// TIA Portal project "TIA_V16_ScalingFunctionExample" (V16)

(* hardware
DEVICE "S71500/ET200MP station_1"  S7-1500 station
   slot 0: "Rail_0"  Rack  6ES7 590-1***0-0AA0
   slot 0: "PS 25W 24VDC_1"  PS 25W 24VDC  6ES7 505-0KA00-0AB0  V1.0
   slot 1: "PLC_1"  CPU 1511F-1 PN  6ES7 511-1FK01-0AB0  V1.8
   slot 2: "DI 16x24VDC HF_1"  DI 16x24VDC HF  6ES7 521-1BH00-0AB0  V2.0
   slot 3: "DQ 16x24VDC/0.5A ST_1"  DQ 16x24VDC/0.5A ST  6ES7 522-1BH00-0AB0  V2.0
   slot 4: "AI 4xU/I/RTD/TC ST_1"  AI 4xU/I/RTD/TC ST  6ES7 531-7QD00-0AB0  V1.0
   slot 5: "AQ 4xU/I ST_1"  AQ 4xU/I ST  6ES7 532-5HD00-0AB0  V2.0
DEVICE "SCALANCE X005"  SCALANCE X-Station
   slot 0: "SCALANCE X rack"  Rail
   slot 0: "Switch_1"  6GK5 005-0BA00-1AA3  V1.0
DEVICE "HMI_1"  TP1200 Comfort
   slot 0: "HMI_1"  TP1200 Comfort  6AV2 124-0MC01-0AX0  16.0.0.0
   slot 1: "HMI_RT_1"  TP1200 Comfort  6AV2 124-0MC01-0AX0  16.0.0.0
   slot 5: "HMI_1.IE_CP_1"  PROFINET Interface  16.0.0.0
      slot 1: "PROFINET Interface_1"  PROFINET Interface
         slot 1: "Port_1"  Port
         slot 2: "Port_2"  Port
   slot 7: "HMI_1.MPI/DP_CP_1"  MPI/DP Interface  16.0.0.0
*)

// ===== PLC "PLC_1"  CPU 1511F-1 PN =====
// protected blocks, not shown: "Main_Safety_RTG1_1", "Main_Safety_RTG1_DB_1"

TYPE "Data Exchange"
TITLE = Data Exchange Between Working Areas
VERSION : 0.1
   STRUCT
      "Working Area 1 Completed" : Bool;
      "Working Area 1 Can Work" : Bool;
      "Working Area 1 Can't Work" : Bool;
      "Working Area 2 Completed" : Bool;
      "Working Area 2 Can Work" : Bool;
      "Working Area 2 Can't  Work" : Bool;
      "Working Area 3 Completed" : Bool;
      "Working Area 3 Can Work" : Bool;
      "Working Area 3 Can't Work" : Bool;
      "Working Area 4 Completed" : Bool;
      "Working Area 4 Can Work" : Bool;
      "Working Area 4 Can't Work" : Bool;
      "WA2 Proof Station OK" : Bool;
      "WA2 Proof Station NOk" : Bool;
      "WA3 Ignition OK" : Bool;
      "WA3 Ignition NOK" : Bool;
      "WA3 Chamber Pressure OK" : Bool;
      "WA3 Chamber Pressure NOK" : Bool;
      Spare1 : Bool;
      Spare2 : Bool;
      Spare3 : Bool;
      Spare4 : Bool;
      Spare5 : Bool;
      Spare6 : Bool;
      Spare7 : Bool;
      Spare8 : Bool;
      Spare9 : Bool;
      Spare10 : Bool;
      Spare11 : Bool;
      Spare12 : Bool;
      Spare13 : Bool;
      Spare14 : Bool;
      Element_1 : Int;
      Element_2 : Int;
      Element_3 : Int;
      Element_4 : Int;
      Element_5 : Int;
      Element_6 : Real;
      Element_8 : Real;
      Element_7 : Real;
      Element_9 : Real;
      Element_10 : Real;
      Rec_PartID : Int;   // Part Record ID Number / 记录ID号
      Rec_Dose_Setting : DInt;   // record recipe dosing setting / 充气设置
      Rec_Gas_Setting_1 : Real;   // record recipe gas setting for shot 1
      Rec_O2_Setting_1 : Real;   // record recipe O2 setting for shot 2
      Rec_Part_Qty : Int;   // record part fixture quanity / 夹具数量
      Rec_Part_weight : Real;   // record recipe part weight
      Rec_shot_type : Int;   // Record recipe shot type
      Rec_Part_image : Array[1..14] of Char;   // PLC part image
      Rec_Fixture_Ref : Array[1..14] of Char;   // record part fixture reference / 夹具参考
      Rec_Part_material : Array[1..14] of Char;   // record part material / 零件材料
      Rec_Part_Name : Array[1..14] of Char;   // record name of part / 记录名称
      Rec_Part_Ref : String[14] := '0';   // record part reference / 零件参考
      Rec_Mix_type1 : Bool;   // record recipe mix type
      Rec_Gas_Setting_2 : Real;   // record recipe gas setting for shot 2
      Rec_O2_Setting_2 : Real;   // record recipe O2 setting for shot 2
      Val_Calibrated_Gas : Int;
      Val_Calibrated_O2 : Int;
      Val_Cailbrated_Gas_Upper : Int;
      Val_Calibrated_Gas_Lower : Int;
      Val_Calibrated_O2_Upper : Int;
      Val_Calibrated_O2_Lower : Int;
      Val_Setting_Gas_Shot_1 : Int;   // Value sent to analog controller for output / 输出值
      Val_Setting_Gas_Shot_2 : Int;   // Value sent to analog controller for output / 输出值
      Val_Setting_O2_Shot_1 : Int := 750;   // Value sent to analog controller for output / 输出值
      Val_Setting_O2_Shot_2 : Int;   // Value sent to analog controller for output / 输出值
      Dose_Setting_Applied : DInt;   // Dosing Stroke Value Applied to Cycle
      BAR_CODE : String[20];
      Rec_MFC_Gas_Setpoint : DInt;
      Rec_MFC_O2_Setpoint : DInt;
   END_STRUCT;
   // Rec_Part_image[1] := '0';
   // Rec_Fixture_Ref[1] := '0';
   // Rec_Part_material[1] := '0';
   // Rec_Part_Name[1] := '0';
END_TYPE

TYPE "UDT_ScalingInputOutput"
   STRUCT
      IN_PV : Word;   // input process value
      IN_OUT_VAL_MIN : Real;   // output value Low limit
      IN_OUT_VAL_MAX : Real;   // output value High limit
      IN_MIN : Real;   // input value Low limit
      IN_MAX : Real;   // input value High limit
      OUT_VAL : Real;   // Output scaled signal
   END_STRUCT;
END_TYPE

TYPE "UDT_ValveActiveConditions_Type_A001"
   STRUCT
      ConditionA : Bool;
      ConditionB : Bool;
      ConditionC : Bool;
   END_STRUCT;
END_TYPE

TYPE "UDT_ValveActiveConditions_Type_A002"
   STRUCT
      ConditionA : Bool;
      ConditionB : Bool;
   END_STRUCT;
END_TYPE

TYPE "UDT_ScalingInput"
   STRUCT
      IN_PV : Word;   // input process value
      IN_OUT_VAL_MIN : Real;   // output value Low limit
      IN_OUT_VAL_MAX : Real;   // output value High limit
      IN_MIN : Real;   // input value Low limit
      IN_MAX : Real;   // input value High limit
   END_STRUCT;
END_TYPE

TYPE "UDT_ScalingOutput"
   STRUCT
      OUT_VAL : Real;   // Output scaled signal
   END_STRUCT;
END_TYPE

// folder: 101_Group_01

DATA_BLOCK "101_DB_ValvesControl"   // DB101
TITLE = 101_DB_Calc_WarmUp_Dosing
{ S7_Optimized_Access := 'FALSE' }
AUTHOR : Jamal
VERSION : 0.1
   VAR
      Valve_1001_Inputs : "UDT_ScalingInput";
      Valve_1001_Outputs : "UDT_ScalingOutput";
      Valve_1002_Inputs : "UDT_ScalingInput";
      Valve_1002_Outputs : "UDT_ScalingOutput";
      Valve_1003_Inputs : "UDT_ScalingInput";
      Valve_1003_Outputs : "UDT_ScalingOutput";
      Valve_1004_Inputs : "UDT_ScalingInput";
      Valve_1004_Outputs : "UDT_ScalingOutput";
      Valve_1001_ActiveConditions : "UDT_ValveActiveConditions_Type_A001";
      LOC_1001_Temperature : Real;
      LOC_1001_Temperature_HighLimit : Real;
      LOC_1001_Temperature_LowLimit : Real;
      Valve_1002_ActiveConditions : "UDT_ValveActiveConditions_Type_A001";
      LOC_1002_Temperature : Real;
      LOC_1002_Temperature_HighLimit : Real;
      LOC_1002_Temperature_LowLimit : Real;
      Valve_1003_ActiveConditions : "UDT_ValveActiveConditions_Type_A002";
      LOC_1003_Temperature : Real;
      LOC_1003_Temperature_HighLimit : Real;
      LOC_1003_Temperature_LowLimit : Real;
      Valve_1004_ActiveConditions : "UDT_ValveActiveConditions_Type_A001";
      LOC_1004_Temperature : Real;
      LOC_1004_Temperature_HighLimit : Real;
      LOC_1004_Temperature_LowLimit : Real;
      HMI : Struct
         ValveSelection : UInt;
         TemperatureSimInput : Word;
         PVSimInput : Word;
         SimOUT_VAL : Real;
         PV_IN_MAX : UInt;
      END_STRUCT;
   END_VAR
BEGIN
END_DATA_BLOCK

// folder: (top level)

ORGANIZATION_BLOCK "Main"   // OB1, LAD, ProgramCycle
TITLE = "Main Program Sweep (Cycle)"
{ S7_Optimized_Access := 'TRUE' }
VERSION : 0.1
   VAR_INPUT
      Initial_Call : Bool;   // Initial call of this OB
      Remanence : Bool;   // =True, if remanent data are available
   END_VAR
   VAR_TEMP
      "Abort_with_SS (Auto to Manual)" : Bool;
      "Abort_with_SS (Manual to Auto)" : Bool;
      Initialize_Graph_Manual_Cycle : Bool;
      Abort_Cycle_Common_bit : Bool;
      TX_Recipe_Transfer : Bool;
      Blk_Return_P1 : Int;
      Blk_Return_P2 : Int;
      Blk_Return_P3 : Int;
      Blk_Return_P4 : Int;
      Blk_Return_P5 : Int;
      Blk_Return_P6 : Int;
      Blk_Return_P7 : Int;
      Blk_Return_P8 : Int;
      Blk_Return_P9 : Int;
   END_VAR
BEGIN

REGION Network 1
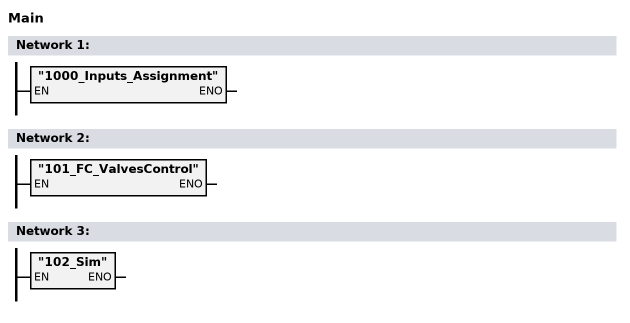
   RUNG wire#powerrail
      "1000_Inputs_Assignment"()
   END_RUNG
   // the same network as SCL:
   "1000_Inputs_Assignment"();
END_REGION

REGION Network 2
   RUNG wire#powerrail
      "101_FC_ValvesControl"()
   END_RUNG
   // the same network as SCL:
   "101_FC_ValvesControl"();
END_REGION

REGION Network 3
   RUNG wire#powerrail
      "102_Sim"()
   END_RUNG
   // the same network as SCL:
   "102_Sim"();
END_REGION
END_ORGANIZATION_BLOCK

// folder: 100_General

FUNCTION "200_ValveControl_Type_A001" : Void   // FC200, SCL
TITLE = 200_ValveControl_Type_A001
{ S7_Optimized_Access := 'TRUE' }
VERSION : 0.1
   VAR_INPUT
      Inputs : "UDT_ScalingInput";
      OUT_VAL_FullOpen : Bool;
      Temperature : Real;
      Temperature_HighLimit : Real;
      Temperature_LowLimit : Real;
      Valve_ActiveConditions : "UDT_ValveActiveConditions_Type_A001";
   END_VAR
   VAR_OUTPUT
      Outputs : "UDT_ScalingOutput";
   END_VAR
BEGIN

   (* Valve_Type_A001 *)

   IF #Temperature >=#Temperature_HighLimit AND #OUT_VAL_FullOpen THEN
       #Outputs.OUT_VAL := 100;
   ELSIF #Temperature >=#Temperature_HighLimit AND NOT #OUT_VAL_FullOpen THEN
       #Outputs.OUT_VAL := #Inputs.IN_OUT_VAL_MAX;
   ELSIF #Temperature >#Temperature_LowLimit AND #Temperature <#Temperature_HighLimit THEN
       "Scaling_Function_1"(IN_PV := #Inputs.IN_PV,
                            IN_OUT_VAL_MIN := #Inputs.IN_OUT_VAL_MIN,
                            IN_OUT_VAL_MAX := #Inputs.IN_OUT_VAL_MAX,
                            IN_MIN := #Inputs.IN_MIN,
                            IN_MAX := #Inputs.IN_MAX,
                            OUT_VAL => #Outputs.OUT_VAL);
   ELSIF #Temperature <=#Temperature_LowLimit THEN
       #Outputs.OUT_VAL := 0;
   END_IF;

   IF NOT #Valve_ActiveConditions.ConditionA OR NOT #Valve_ActiveConditions.ConditionB OR NOT #Valve_ActiveConditions.ConditionC THEN
       #Outputs.OUT_VAL := 0;
   END_IF;
END_FUNCTION

FUNCTION "201_ValveControl_Type_A002" : Void   // FC201, SCL
TITLE = 200_ValveControl_Type_A001
{ S7_Optimized_Access := 'TRUE' }
VERSION : 0.1
   VAR_INPUT
      Inputs : "UDT_ScalingInput";
      OUT_VAL_FullOpen : Bool;
      Temperature : Real;
      Temperature_HighLimit : Real;
      Temperature_LowLimit : Real;
      Valve_ActiveConditions : "UDT_ValveActiveConditions_Type_A002";
   END_VAR
   VAR_OUTPUT
      Outputs : "UDT_ScalingOutput";
   END_VAR
BEGIN

   (* Valve_Type_A002 *)

   IF #Temperature >=#Temperature_HighLimit AND #OUT_VAL_FullOpen THEN
       #Outputs.OUT_VAL := 100;
   ELSIF #Temperature >=#Temperature_HighLimit AND NOT #OUT_VAL_FullOpen THEN
       #Outputs.OUT_VAL := #Inputs.IN_OUT_VAL_MAX;
   ELSIF #Temperature >#Temperature_LowLimit AND #Temperature <#Temperature_HighLimit THEN
       "Scaling_Function_1"(IN_PV := #Inputs.IN_PV,
                            IN_OUT_VAL_MIN := #Inputs.IN_OUT_VAL_MIN,
                            IN_OUT_VAL_MAX := #Inputs.IN_OUT_VAL_MAX,
                            IN_MIN := #Inputs.IN_MIN,
                            IN_MAX := #Inputs.IN_MAX,
                            OUT_VAL => #Outputs.OUT_VAL);
   ELSIF #Temperature <=#Temperature_LowLimit THEN
       #Outputs.OUT_VAL := 0;
   END_IF;

   IF NOT #Valve_ActiveConditions.ConditionA OR NOT #Valve_ActiveConditions.ConditionB THEN
       #Outputs.OUT_VAL := 0;
   END_IF;
END_FUNCTION

FUNCTION "Scaling_Function_1" : Void   // FC700, SCL
TITLE = ScalingOut_0_10V
{ S7_Optimized_Access := 'TRUE' }
AUTHOR : Jamal
VERSION : 0.1
   VAR_INPUT
      IN_PV : Word;   // input process value
      IN_OUT_VAL_MIN : Real;   // output value Low limit
      IN_OUT_VAL_MAX : Real;   // output value High limit
      IN_MIN : Real;   // input value Low limit
      IN_MAX : Real;   // input value High limit
   END_VAR
   VAR_OUTPUT
      OUT_VAL : Real;   // output scaled signal
   END_VAR
BEGIN
   (*
   //JMu_26.09.2019
   IN_OUT_VAL_MIN = output value Low limit
   IN_OUT_VAL_MAX = output value High limit
   //Output value High Limit & Low Limit (this is what you want or in case of standard 0-10V/4-20mA actuators its IN_OUT_VAL_MIN=0 & IN_OUT_VAL_MAX=27648).
   //In case if we want a valve to Open 30% (27648X30%=8294.4) from very first actuation then IN_OUT_VAL_MIN=8294.4 & IN_OUT_VAL_MAX=27648 

   IN_MIN = input value Low limit
   IN_MAX = input value High limit
   //In case of standard 0-10V/4-20mA sensors the values are IN_MIN=0 & IN_MAX=27648 or 32000.
   //In case if we want to scale an inside variable value e.g Temperature in Deg Centigrade(0°-65°Cen) then IN_MIN=0 & IN_MAX=65. 

   *)

   #OUT_VAL := (#IN_OUT_VAL_MAX - #IN_OUT_VAL_MIN) / (#IN_MAX - #IN_MIN) * (#IN_PV - #IN_MIN) + #IN_OUT_VAL_MIN;
END_FUNCTION

FUNCTION "Scaling_Function_2" : Void   // FC701, FBD
TITLE = Scaling_Function_2
{ S7_Optimized_Access := 'TRUE' }
VERSION : 0.1
   VAR_INPUT
      Input_Min : Int;
      Input_Max : Int;
      Input_PV : Int;
      Output_Min : Real;
      Output_Max : Real;
   END_VAR
   VAR_OUTPUT
      SV : Real;
   END_VAR
   VAR_TEMP
      tv : Real;
   END_VAR
BEGIN

REGION Network 1
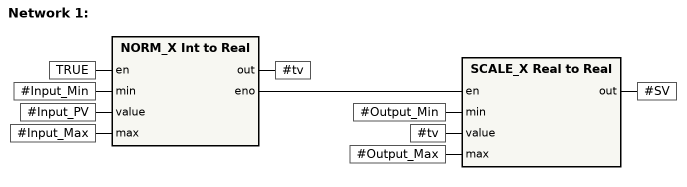
   IF TRUE THEN
       #tv := NORM_X(MIN := #Input_Min, VALUE := #Input_PV, MAX := #Input_Max);
       #SV := SCALE_X(MIN := #Output_Min, VALUE := #tv, MAX := #Output_Max);
   END_IF;
END_REGION
END_FUNCTION

// folder: 101_Group_01

FUNCTION "101_FC_ValvesControl" : Void   // FC101, SCL
{ S7_Optimized_Access := 'TRUE' }
VERSION : 0.1
BEGIN
   (* Scaling outputs for all 4 valves *)
   //Valve_1001/TypeA001
   //input in between min 0 - max 27648 
   //output needs to be in between min 0% - max 80%
   "200_ValveControl_Type_A001"(Inputs := "101_DB_ValvesControl".Valve_1001_Inputs,
                                OUT_VAL_FullOpen := FALSE,
                                Temperature := "101_DB_ValvesControl".LOC_1001_Temperature,
                                Temperature_HighLimit := "101_DB_ValvesControl".LOC_1001_Temperature_HighLimit,
                                Temperature_LowLimit := "101_DB_ValvesControl".LOC_1001_Temperature_LowLimit,
                                Valve_ActiveConditions := "101_DB_ValvesControl".Valve_1001_ActiveConditions,
                                Outputs => "101_DB_ValvesControl".Valve_1001_Outputs);


   //Valve_1002/TypeA001
   //input in between min 0 - max 27648
   //output needs to be in between min 0% - max 70%
   "200_ValveControl_Type_A001"(Inputs := "101_DB_ValvesControl".Valve_1002_Inputs,
                                OUT_VAL_FullOpen := FALSE,
                                Temperature := "101_DB_ValvesControl".LOC_1002_Temperature,
                                Temperature_HighLimit := "101_DB_ValvesControl".LOC_1002_Temperature_HighLimit,
                                Temperature_LowLimit := "101_DB_ValvesControl".LOC_1002_Temperature_LowLimit,
                                Valve_ActiveConditions := "101_DB_ValvesControl".Valve_1002_ActiveConditions,
                                Outputs => "101_DB_ValvesControl".Valve_1002_Outputs);

   //Valve_1003/TypeA002
   //input in between min 0 - max 32000 
   //output needs to be in between min 0% - max 90%
   //when temperature > 69 deg Cen. then OUT_VAL:=100% 
   "201_ValveControl_Type_A002"(Inputs := "101_DB_ValvesControl".Valve_1003_Inputs,
                                OUT_VAL_FullOpen := TRUE,
                                Temperature := "101_DB_ValvesControl".LOC_1003_Temperature,
                                Temperature_HighLimit := "101_DB_ValvesControl".LOC_1003_Temperature_HighLimit,
                                Temperature_LowLimit := "101_DB_ValvesControl".LOC_1003_Temperature_LowLimit,
                                Valve_ActiveConditions := "101_DB_ValvesControl".Valve_1003_ActiveConditions,
                                Outputs => "101_DB_ValvesControl".Valve_1003_Outputs);

   //Valve_1004/TypeA001
   //input in between min 0 - max 27648 
   //output needs to be in between min 0% - max 60%
   "200_ValveControl_Type_A001"(Inputs := "101_DB_ValvesControl".Valve_1004_Inputs,
                                OUT_VAL_FullOpen := FALSE,
                                Temperature := "101_DB_ValvesControl".LOC_1004_Temperature,
                                Temperature_HighLimit := "101_DB_ValvesControl".LOC_1004_Temperature_HighLimit,
                                Temperature_LowLimit := "101_DB_ValvesControl".LOC_1004_Temperature_LowLimit,
                                Valve_ActiveConditions := "101_DB_ValvesControl".Valve_1004_ActiveConditions,
                                Outputs => "101_DB_ValvesControl".Valve_1004_Outputs);


   //HMI variables
END_FUNCTION

FUNCTION "102_Sim" : Void   // FC102, SCL
TITLE = 102_Sim
{ S7_Optimized_Access := 'TRUE' }
VERSION : 0.1
BEGIN

   IF "101_DB_ValvesControl".HMI.ValveSelection = 1 THEN
       "101_DB_ValvesControl".Valve_1001_Inputs.IN_PV := "101_DB_ValvesControl".HMI.PVSimInput;
       "101_DB_ValvesControl".LOC_1001_Temperature := WORD_TO_INT("101_DB_ValvesControl".HMI.TemperatureSimInput);
       "101_DB_ValvesControl".HMI.SimOUT_VAL := "101_DB_ValvesControl".Valve_1001_Outputs.OUT_VAL;
       "101_DB_ValvesControl".HMI.PV_IN_MAX := 27648;
   ELSIF "101_DB_ValvesControl".HMI.ValveSelection = 2 THEN
       "101_DB_ValvesControl".Valve_1002_Inputs.IN_PV := "101_DB_ValvesControl".HMI.PVSimInput;
       "101_DB_ValvesControl".LOC_1002_Temperature := WORD_TO_INT("101_DB_ValvesControl".HMI.TemperatureSimInput);
       "101_DB_ValvesControl".HMI.SimOUT_VAL := "101_DB_ValvesControl".Valve_1002_Outputs.OUT_VAL;
       "101_DB_ValvesControl".HMI.PV_IN_MAX := 27648;
   ELSIF "101_DB_ValvesControl".HMI.ValveSelection = 3 THEN
       "101_DB_ValvesControl".Valve_1003_Inputs.IN_PV := "101_DB_ValvesControl".HMI.PVSimInput;
       "101_DB_ValvesControl".LOC_1003_Temperature := WORD_TO_INT("101_DB_ValvesControl".HMI.TemperatureSimInput);
       "101_DB_ValvesControl".HMI.SimOUT_VAL := "101_DB_ValvesControl".Valve_1003_Outputs.OUT_VAL;
       "101_DB_ValvesControl".HMI.PV_IN_MAX := 32000;
   ELSIF "101_DB_ValvesControl".HMI.ValveSelection = 4 THEN
       "101_DB_ValvesControl".Valve_1004_Inputs.IN_PV := "101_DB_ValvesControl".HMI.PVSimInput;
       "101_DB_ValvesControl".LOC_1004_Temperature := WORD_TO_INT("101_DB_ValvesControl".HMI.TemperatureSimInput);
       "101_DB_ValvesControl".HMI.SimOUT_VAL := "101_DB_ValvesControl".Valve_1004_Outputs.OUT_VAL;
       "101_DB_ValvesControl".HMI.PV_IN_MAX := 27648;
   END_IF;
END_FUNCTION

FUNCTION "1000_Inputs_Assignment" : Void   // FC1000, SCL
TITLE = 1000_Input_Assignment
{ S7_Optimized_Access := 'TRUE' }
VERSION : 0.1
BEGIN
   "101_DB_ValvesControl".Valve_1001_Inputs.IN_MIN := 0;
   "101_DB_ValvesControl".Valve_1001_Inputs.IN_MAX := 27648;
   "101_DB_ValvesControl".Valve_1001_Inputs.IN_OUT_VAL_MIN := 0;
   "101_DB_ValvesControl".Valve_1001_Inputs.IN_OUT_VAL_MAX := 80;
   "101_DB_ValvesControl".LOC_1001_Temperature_HighLimit := 69;
   "101_DB_ValvesControl".LOC_1001_Temperature_LowLimit := 17;
   "101_DB_ValvesControl".Valve_1001_ActiveConditions.ConditionA := TRUE;
   "101_DB_ValvesControl".Valve_1001_ActiveConditions.ConditionB := TRUE;
   "101_DB_ValvesControl".Valve_1001_ActiveConditions.ConditionC := TRUE;

   "101_DB_ValvesControl".Valve_1002_Inputs.IN_MIN := 0;
   "101_DB_ValvesControl".Valve_1002_Inputs.IN_MAX := 27648;
   "101_DB_ValvesControl".Valve_1002_Inputs.IN_OUT_VAL_MIN := 0;
   "101_DB_ValvesControl".Valve_1002_Inputs.IN_OUT_VAL_MAX := 60;
   "101_DB_ValvesControl".LOC_1002_Temperature_HighLimit := 69;
   "101_DB_ValvesControl".LOC_1002_Temperature_LowLimit := 17;
   "101_DB_ValvesControl".Valve_1002_ActiveConditions.ConditionA := TRUE;
   "101_DB_ValvesControl".Valve_1002_ActiveConditions.ConditionB := TRUE;
   "101_DB_ValvesControl".Valve_1002_ActiveConditions.ConditionC := TRUE;

   "101_DB_ValvesControl".Valve_1003_Inputs.IN_MIN := 0;
   "101_DB_ValvesControl".Valve_1003_Inputs.IN_MAX := 32000;
   "101_DB_ValvesControl".Valve_1003_Inputs.IN_OUT_VAL_MIN := 0;
   "101_DB_ValvesControl".Valve_1003_Inputs.IN_OUT_VAL_MAX := 90;
   "101_DB_ValvesControl".LOC_1003_Temperature_HighLimit := 69;
   "101_DB_ValvesControl".LOC_1003_Temperature_LowLimit := 17;
   "101_DB_ValvesControl".Valve_1003_ActiveConditions.ConditionA := TRUE;
   "101_DB_ValvesControl".Valve_1003_ActiveConditions.ConditionB := TRUE;

   "101_DB_ValvesControl".Valve_1004_Inputs.IN_MIN := 0;
   "101_DB_ValvesControl".Valve_1004_Inputs.IN_MAX := 27648;
   "101_DB_ValvesControl".Valve_1004_Inputs.IN_OUT_VAL_MIN := 0;
   "101_DB_ValvesControl".Valve_1004_Inputs.IN_OUT_VAL_MAX := 60;
   "101_DB_ValvesControl".LOC_1004_Temperature_HighLimit := 69;
   "101_DB_ValvesControl".LOC_1004_Temperature_LowLimit := 17;
   "101_DB_ValvesControl".Valve_1004_ActiveConditions.ConditionA := TRUE;
   "101_DB_ValvesControl".Valve_1004_ActiveConditions.ConditionB := TRUE;
   "101_DB_ValvesControl".Valve_1004_ActiveConditions.ConditionC := TRUE;
END_FUNCTION

FUNCTION "2000_Outputs_Assignment" : Void   // FC2000, SCL
TITLE = 2000_Output_Assignment
{ S7_Optimized_Access := 'TRUE' }
VERSION : 0.1
BEGIN
END_FUNCTION

(* ===== HMI "HMI_RT_1" =====
system functions are stored by id; their names below are inferred from use
connection "HMI_Connection_1": ETHERNET, S7_1500_OMS

HMI tags "Default tag table"
   "Tag_ScreenNumber" : UInt, internal
   "101_DB_ValvesControl_HMI_ValveSelection" : UInt = PLC "101_DB_ValvesControl".HMI.ValveSelection AT %DB101.DBW144, 1 s
   "101_DB_ValvesControl_HMI_PVSimInput" : Word = PLC "101_DB_ValvesControl".HMI.PVSimInput AT %DB101.DBW148, 1 s
   "101_DB_ValvesControl_HMI_Temperature" : Word = PLC "101_DB_ValvesControl".HMI.TemperatureSimInput AT %DB101.DBW146, 1 s
   "101_DB_ValvesControl_HMI_SimOUT_VAL" : Real = PLC "101_DB_ValvesControl".HMI.SimOUT_VAL AT %DB101.DBD150, 1 s
   "101_DB_ValvesControl_HMI_PV_IN_MAX" : UInt = PLC "101_DB_ValvesControl".HMI.PV_IN_MAX AT %DB101.DBW154, 1 s

text list "ValveSelection": 1 'Valve 1001'; 2 'Valve 1002'; 3 'Valve 1003'; 4 'Valve 1004'

screen "Root screen" 1280x740, template "Template_1"
   on GenerateScreen: SetTag("Tag_ScreenNumber", 1)
   TextField "HmiScreenItemData" at 58,39 size 191x27; Text 'PV / Willkommen zum HMI_1 (TP1200 Comfort)!'
   TextField "HmiScreenItemData_1" at 39,143 size 214x27; Text 'Temperature / Willkommen zum HMI_1 (TP1200 Comfort)!'
   Slider "Slider_1" at 257,19 size 803x61; Caption 'SIMATIC'
      ProcessValue <- "101_DB_ValvesControl_HMI_PVSimInput"
      MaximumValue <- "101_DB_ValvesControl_HMI_PV_IN_MAX"
   Slider "Slider_2" at 257,133 size 803x61; Caption 'SIMATIC'
      ProcessValue <- "101_DB_ValvesControl_HMI_Temperature"
   TrendView "Trend view_1" at 36,259 size 1213x408
   SymbolicIOField "Symbolic I/O field_1" at 1078,209 size 170x42; TextOff '0'; TextOn '1'; TextList "ValveSelection"
      ProcessValue <- "101_DB_ValvesControl_HMI_ValveSelection"
   TextField "Text field_1" at 1073,184 size 148x25; Text 'Valve selection'

Template "Template_1" 1280x740
   Button "Exit" at 1200,679 size 78x59; TextOff 'Exit / Beenden'; PictureOff "ExitRuntime_TP1200_Comfort_TR"; PictureOn "ExitRuntime_TP1200_Comfort_TR"
      on Release: StopRuntime(0)
   Button "Template_Button" at 1120,679 size 78x59; TextOff 'Text'
   Button "Template_Button_1" at 1040,679 size 78x59; TextOff 'Text'
   Button "Template_Button_2" at 960,679 size 78x59; TextOff 'Text'
   Button "Template_Button_3" at 880,679 size 78x59; TextOff 'Text'
   Button "Template_Button_4" at 800,679 size 78x59; TextOff 'Text'
   Button "Template_Button_5" at 720,679 size 78x59; TextOff 'Text'
   Button "Template_Button_6" at 640,679 size 78x59; TextOff 'Text'
   Button "Template_Button_7" at 561,679 size 78x59; TextOff 'Text'
   Button "Template_Button_8" at 481,679 size 78x59; TextOff 'Text'
   Button "Template_Button_9" at 401,679 size 78x59; TextOff 'Text'
   Button "Template_Button_10" at 321,679 size 78x59; TextOff 'Text'
   Button "Template_Button_11" at 241,679 size 78x59; TextOff 'Text'
   Button "Template_Button_12" at 161,679 size 78x59; TextOff 'Text'
   Button "Alarms" at 81,679 size 78x59; TextOff 'Alarms / Meldungen'; PictureOff "AlarmDisplay_TP1200_Comfort_TR"; PictureOn "AlarmDisplay_TP1200_Comfort_TR"
      on Release: function_ef3f5d25("Alarm window_Unacknowledged", -1)
   Button "Start screen" at 1,679 size 78x59; TextOff 'Start screen / Startbild'; PictureOff "NavigateHome_TP1200_Comfort_TR"; PictureOn "NavigateHome_TP1200_Comfort_TR"
      on Release: ActivateScreen("Root screen", 0)
*)